// TIA Portal project "Lagerregal_5" (V20) (continued)

   IF #"PTRIG_MDB_Z-Neg".Q THEN
       "HMI_Schnittstelle".Kraene.Kran_1.Kran_Pos."Z-Soll" -= UINT_TO_INT("HMI_Schnittstelle".HMI.Inkrement);
   END_IF;
END_REGION
END_FUNCTION_BLOCK

FUNCTION_BLOCK "Ein_HMI"   // FB10, FBD
{ S7_Optimized_Access := 'TRUE' }
VERSION : 0.1
BEGIN
END_FUNCTION_BLOCK

FUNCTION "Meldungen" : Void   // FC10, SCL
{ S7_Optimized_Access := 'TRUE' }
VERSION : 0.1
BEGIN
   // Slice Zugriff programmieren
   // d.h. wir können auf die Einzelbits einer Ganzzahlvariable (INT, DINT, etc.)
   // bzw. einer Bitfolge (Byte, Word, etc.) zugreifen.

   // Bits:        Variable.%X0
   // Bytes:       Variable.%B0
   // Word:        Variable.%W0
   // DWord:       Variable.%D0


   "HMI_Schnittstelle".Bitmeldungen.%X0 := "HMI_Schnittstelle".Eingaenge.S2;
   "HMI_Schnittstelle".Bitmeldungen.%X1 := "HMI_Schnittstelle".Eingaenge.S1;
   "HMI_Schnittstelle".Bitmeldungen.%X2 := "HMI_Schnittstelle".Betriebsart.Hand;
   "HMI_Schnittstelle".Bitmeldungen.%X3 := "HMI_Schnittstelle".Betriebsart.Automatik;
END_FUNCTION

// folder: Kransteuerung

FUNCTION_BLOCK "FC_Kran_beladen"   // FB25, FBD
{ S7_Optimized_Access := 'TRUE' }
VERSION : 0.1
   VAR_INPUT
      "eKran_Z-Ist" : Int;
      eSchrittnummer : Int;
   END_VAR
   VAR_OUTPUT
      aGabel : Bool;
      aBeladen : Bool;
      "aKran_Z-Soll" : Int;
   END_VAR
   VAR
      PTRIG_Schritt2 : Bool;
   END_VAR
   VAR_TEMP   // added for the SCL form of the ladder/FBD networks
      _w1 : Bool;
      _w2 : Bool;
   END_VAR
BEGIN

REGION Network 1: Gabel zur Seite ausfahren
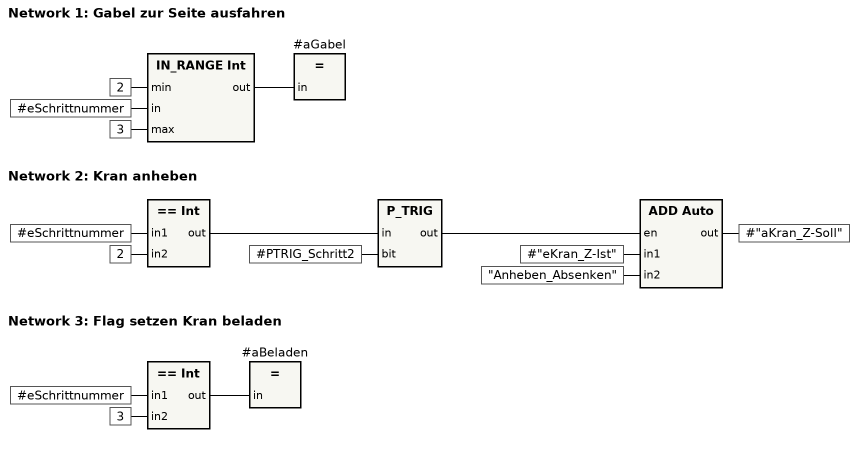
   #aGabel := (2 <= #eSchrittnummer) AND (#eSchrittnummer <= 3);
END_REGION

REGION Network 2: Kran anheben
   #_w1 := #eSchrittnummer = 2;
   #_w2 := #_w1 AND NOT #PTRIG_Schritt2;   // rising edge
   #PTRIG_Schritt2 := #_w1;
   IF #_w2 THEN #"aKran_Z-Soll" := #"eKran_Z-Ist" + "Anheben_Absenken"; END_IF;
END_REGION

REGION Network 3: Flag setzen Kran beladen
   #aBeladen := #eSchrittnummer = 3;
END_REGION
END_FUNCTION_BLOCK

FUNCTION_BLOCK "FC_Kran_entladen"   // FB26, FBD
{ S7_Optimized_Access := 'TRUE' }
VERSION : 0.1
   VAR_INPUT
      "eKran_Z-Ist" : Int;
      eSchrittnummer : Int;
   END_VAR
   VAR_OUTPUT
      aGabel : Bool;
      aBeladen : Bool;
      "aKran_Z-Soll" : Int;
   END_VAR
   VAR
      PTRIG_Schritt2 : Bool;
   END_VAR
   VAR_TEMP   // added for the SCL form of the ladder/FBD networks
      _w1 : Bool;
      _w2 : Bool;
   END_VAR
BEGIN

REGION Network 1: Gabel zur Seite ausfahren
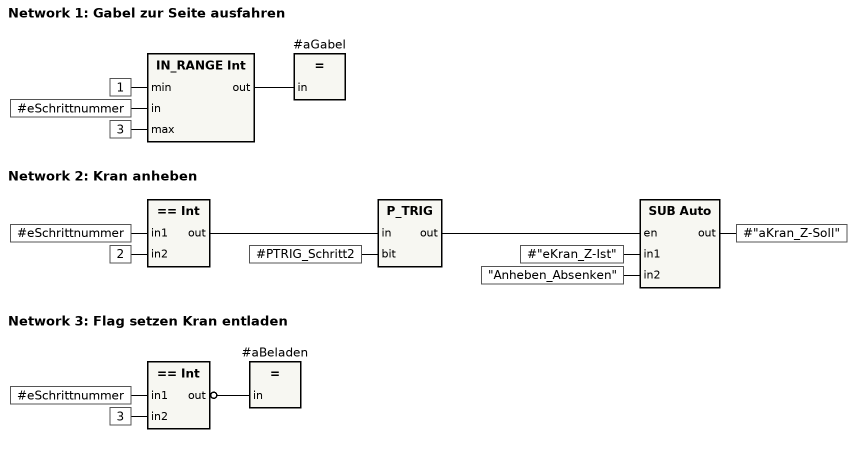
   #aGabel := (1 <= #eSchrittnummer) AND (#eSchrittnummer <= 3);
END_REGION

REGION Network 2: Kran anheben
   #_w1 := #eSchrittnummer = 2;
   #_w2 := #_w1 AND NOT #PTRIG_Schritt2;   // rising edge
   #PTRIG_Schritt2 := #_w1;
   IF #_w2 THEN #"aKran_Z-Soll" := #"eKran_Z-Ist" - "Anheben_Absenken"; END_IF;
END_REGION

REGION Network 3: Flag setzen Kran entladen
   #aBeladen := NOT (#eSchrittnummer = 3);
END_REGION
END_FUNCTION_BLOCK

FUNCTION_BLOCK "Ein_Kran"   // FB30, FBD
{ S7_Optimized_Access := 'TRUE' }
VERSION : 0.1
   VAR
      NTRIG_MDB_1B2 : F_TRIG;
      NTRIG_MDB_2B2 : F_TRIG;
      NTRIG_MDB_5B1 : F_TRIG;
   END_VAR
BEGIN

REGION Network 1 (SCL): Sensoren Kran_1
   "HMI_Schnittstelle".Eingaenge."6B1" := "6B1";
   "HMI_Schnittstelle".Eingaenge."6B2" := "6B2";
   "HMI_Schnittstelle".Eingaenge."6B3" := "6B3";
END_REGION

REGION Network 2: Kran_1 Position einlesen
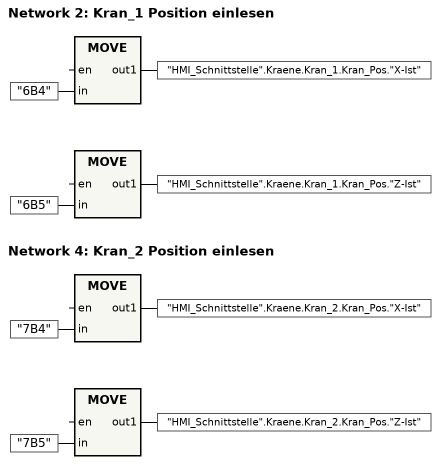
   "HMI_Schnittstelle".Kraene.Kran_1.Kran_Pos."X-Ist" := "6B4";
   "HMI_Schnittstelle".Kraene.Kran_1.Kran_Pos."Z-Ist" := "6B5";
END_REGION

REGION Network 3 (SCL): Sensoren Kran_2
   "HMI_Schnittstelle".Eingaenge."7B1" := "7B1";
   "HMI_Schnittstelle".Eingaenge."7B2" := "7B2";
   "HMI_Schnittstelle".Eingaenge."7B3" := "7B3";
END_REGION

REGION Network 4: Kran_2 Position einlesen
   "HMI_Schnittstelle".Kraene.Kran_2.Kran_Pos."X-Ist" := "7B4";
   "HMI_Schnittstelle".Kraene.Kran_2.Kran_Pos."Z-Ist" := "7B5";
END_REGION
END_FUNCTION_BLOCK

FUNCTION_BLOCK "Prog_Automatik_einlagern"   // FB50, FBD
{ S7_Optimized_Access := 'TRUE' }
VERSION : 0.1
   VAR
      MDB_Schrittkette_einlagern : "Prog_Schrittkette";
      FTRIG_Palette_eingelagert : F_TRIG;
   END_VAR
   VAR_TEMP
      tmpPalette_abgelegt : Int;
      tmpFaecher_durchlaufen : Int;
   END_VAR
BEGIN

REGION Network 1 (SCL): Lagerplatz frei
   IF "HMI_Schnittstelle".Anlagendaten.Fach > 0 AND "HMI_Schnittstelle".Anlagendaten.Fach < 55 THEN
       "HMI_Schnittstelle".Anlagendaten.Regalplatz_frei := "Warenlager".Lager["HMI_Schnittstelle".Anlagendaten.Fach].Bauteil = 0;

       IF NOT "HMI_Schnittstelle".Anlagendaten.Regalplatz_frei AND "HMI_Schnittstelle".Anlagendaten.Fach < 54 THEN
           // Zähle das Fach hoch, wenn das aktuell Fach belegt ist.
           "HMI_Schnittstelle".Anlagendaten.Fach += 1;
       END_IF;
   ELSE
       "HMI_Schnittstelle".Anlagendaten.Regalplatz_frei := FALSE;
   END_IF;


   // Verhindere Endlos-Schleife
   IF #tmpFaecher_durchlaufen = 2 AND NOT "HMI_Schnittstelle".Anlagendaten.Regalplatz_frei THEN
       "HMI_Schnittstelle".Anlagendaten.Fach := 0;
       "HMI_Schnittstelle".Betriebsart.Automatik := FALSE;
   END_IF;
END_REGION

REGION Network 2: Palette abgelegt
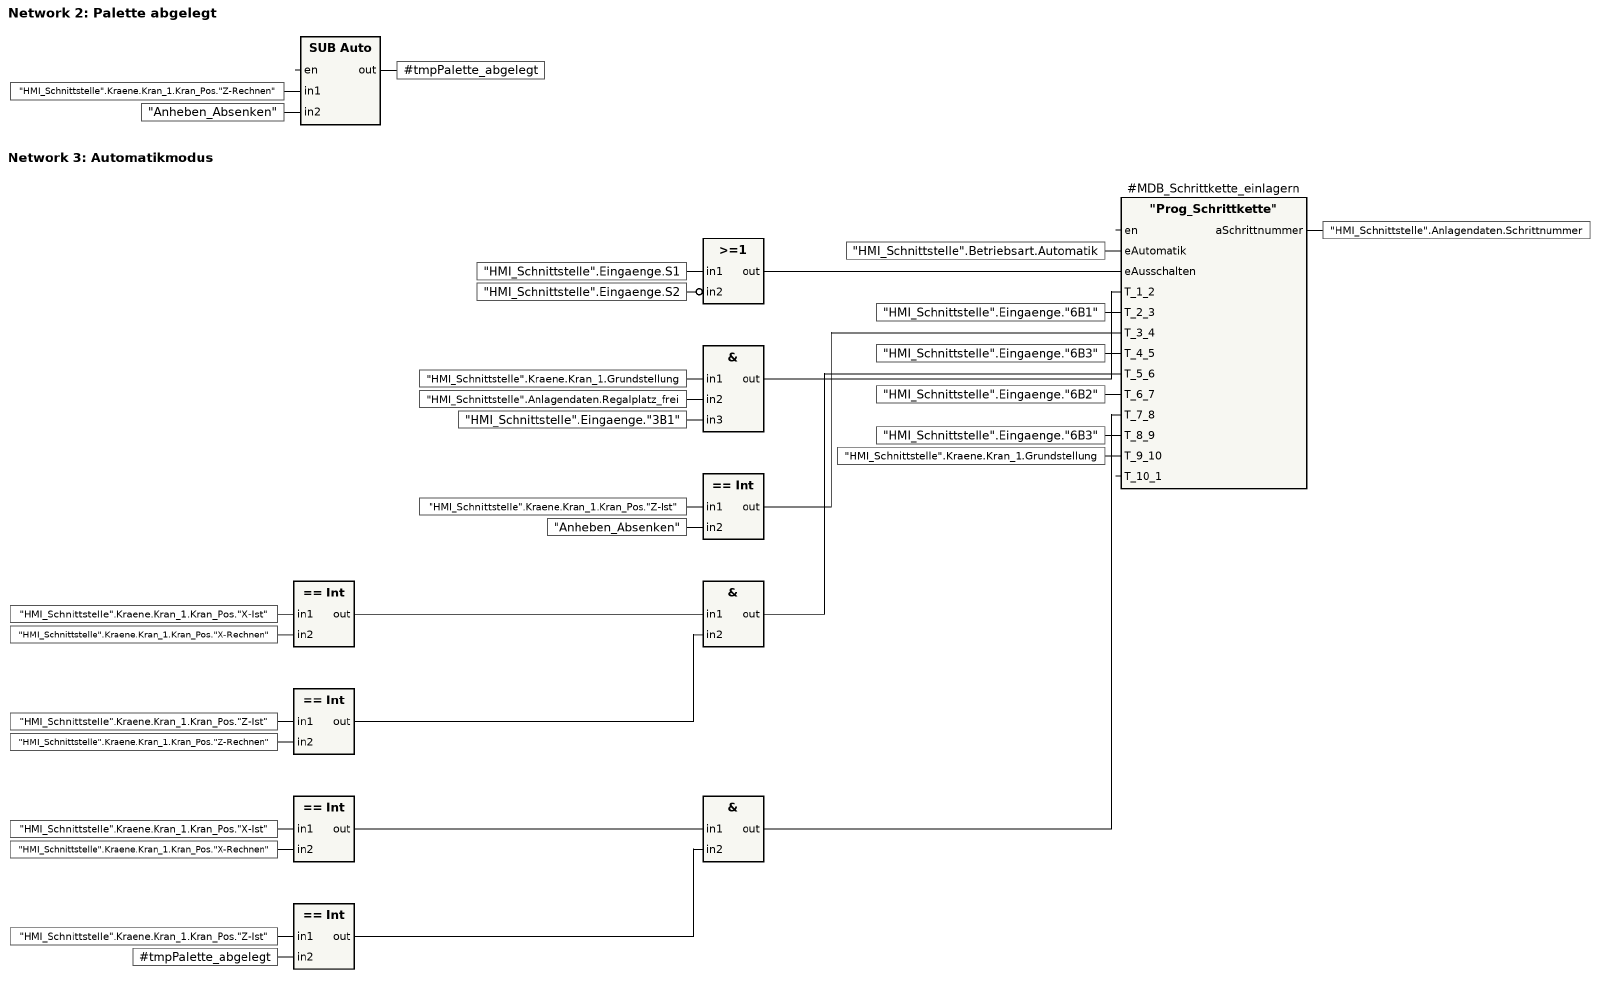
   #tmpPalette_abgelegt := "HMI_Schnittstelle".Kraene.Kran_1.Kran_Pos."Z-Rechnen" - "Anheben_Absenken";
END_REGION

REGION Network 3: Automatikmodus
   #MDB_Schrittkette_einlagern(eAutomatik := "HMI_Schnittstelle".Betriebsart.Automatik,   // "Prog_Schrittkette"
                           eAusschalten := "HMI_Schnittstelle".Eingaenge.S1 OR NOT "HMI_Schnittstelle".Eingaenge.S2,
                           T_1_2 := "HMI_Schnittstelle".Kraene.Kran_1.Grundstellung AND "HMI_Schnittstelle".Anlagendaten.Regalplatz_frei AND "HMI_Schnittstelle".Eingaenge."3B1",
                           T_2_3 := "HMI_Schnittstelle".Eingaenge."6B1",
                           T_3_4 := "HMI_Schnittstelle".Kraene.Kran_1.Kran_Pos."Z-Ist" = "Anheben_Absenken",
                           T_4_5 := "HMI_Schnittstelle".Eingaenge."6B3",
                           T_5_6 := ("HMI_Schnittstelle".Kraene.Kran_1.Kran_Pos."X-Ist" = "HMI_Schnittstelle".Kraene.Kran_1.Kran_Pos."X-Rechnen") AND ("HMI_Schnittstelle".Kraene.Kran_1.Kran_Pos."Z-Ist" = "HMI_Schnittstelle".Kraene.Kran_1.Kran_Pos."Z-Rechnen"),
                           T_6_7 := "HMI_Schnittstelle".Eingaenge."6B2",
                           T_7_8 := ("HMI_Schnittstelle".Kraene.Kran_1.Kran_Pos."X-Ist" = "HMI_Schnittstelle".Kraene.Kran_1.Kran_Pos."X-Rechnen") AND ("HMI_Schnittstelle".Kraene.Kran_1.Kran_Pos."Z-Ist" = #tmpPalette_abgelegt),
                           T_8_9 := "HMI_Schnittstelle".Eingaenge."6B3",
                           T_9_10 := "HMI_Schnittstelle".Kraene.Kran_1.Grundstellung,
                           aSchrittnummer => "HMI_Schnittstelle".Anlagendaten.Schrittnummer);
END_REGION

REGION Network 4 (SCL): Fachnummer erhöhen
   #FTRIG_Palette_eingelagert(CLK := "HMI_Schnittstelle".Anlagendaten.Schrittnummer = 7);


   // Wenn die Palette eingelagert wurde, ...
   IF #FTRIG_Palette_eingelagert.Q THEN
       // ... schreibe die Info über das Bauteil ins Array.
       "Warenlager".Lager["HMI_Schnittstelle".Anlagendaten.Fach].Bauteil := "HMI_Schnittstelle".Anlagendaten.Bauteil;

       // Zähle das Fach hoch und setze das aktuelle Bauteil zurück.
       "HMI_Schnittstelle".Anlagendaten.Fach += 1;
       "HMI_Schnittstelle".Anlagendaten.Bauteil := 0;
   END_IF;

   IF "HMI_Schnittstelle".Anlagendaten.Fach = 54 THEN
       // Setze das Fach 1, wenn am Ende angekommen.
       "HMI_Schnittstelle".Anlagendaten.Fach := 1;
       #tmpFaecher_durchlaufen += 1;
   END_IF;
END_REGION
END_FUNCTION_BLOCK

FUNCTION "Aus_Kran" : Void   // FC30, FBD
{ S7_Optimized_Access := 'TRUE' }
VERSION : 0.1
BEGIN

REGION Network 1 (SCL): Kräne Gabelsteuerung
   "6M1" := "HMI_Schnittstelle".Ausgaenge."6M1";
   "6M2" := "HMI_Schnittstelle".Ausgaenge."6M2";

   "7M1" := "HMI_Schnittstelle".Ausgaenge."7M1";
   "7M2" := "HMI_Schnittstelle".Ausgaenge."7M2";
END_REGION
END_FUNCTION

FUNCTION "FC_Kran_Grundstellung" : Void   // FC31, FBD
{ S7_Optimized_Access := 'TRUE' }
VERSION : 0.1
   VAR_INPUT
      "X-Ist" : Int;
      "Z-Ist" : Int;
      Gabel_mitte : Bool;
   END_VAR
   VAR_OUTPUT
      Heimposition : Bool;
      Grundstellung : Bool;
   END_VAR
BEGIN

REGION Network 1
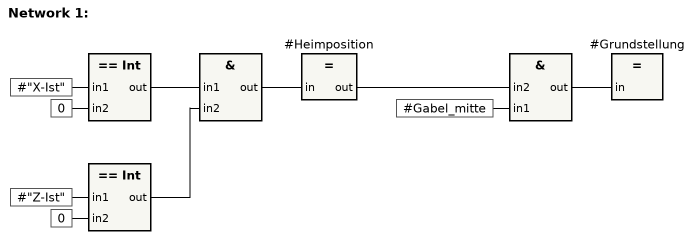
   #Heimposition := (#"X-Ist" = 0) AND (#"Z-Ist" = 0);
   #Grundstellung := #Heimposition AND #Gabel_mitte;
END_REGION
END_FUNCTION

FUNCTION "Staplersteuerung" : Void   // FC70, FBD
{ S7_Optimized_Access := 'TRUE' }
VERSION : 0.1
BEGIN

REGION Network 1: Sollposition X
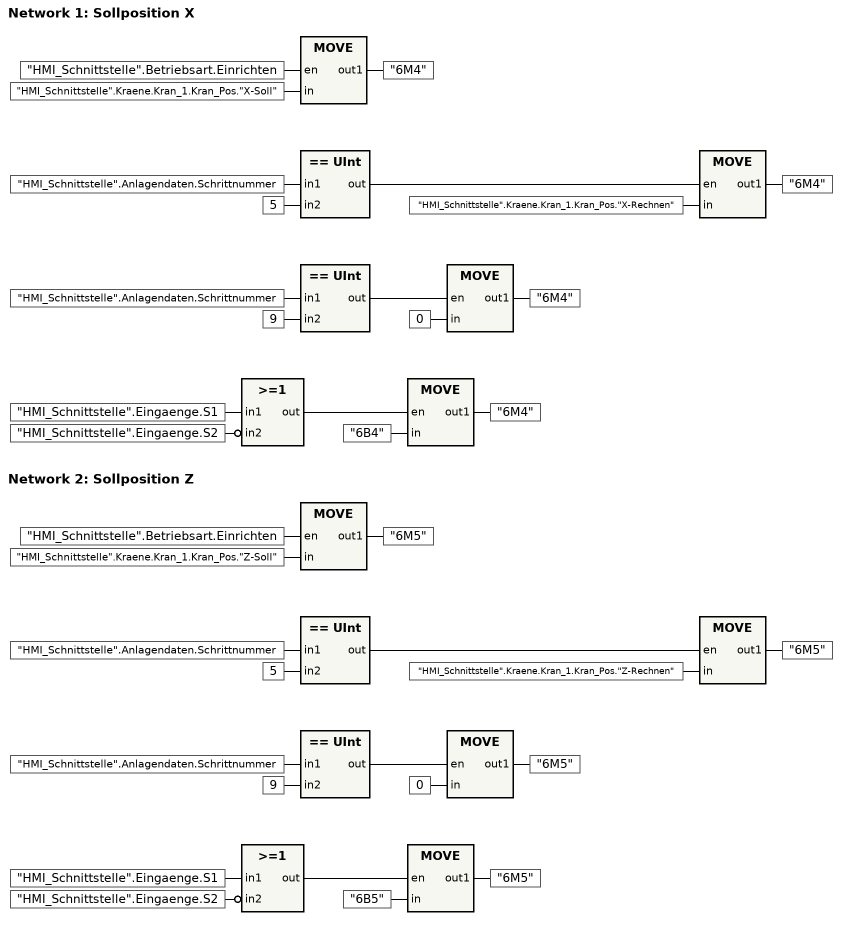
   IF "HMI_Schnittstelle".Betriebsart.Einrichten THEN
       "6M4" := "HMI_Schnittstelle".Kraene.Kran_1.Kran_Pos."X-Soll";
   END_IF;
   IF "HMI_Schnittstelle".Anlagendaten.Schrittnummer = 5 THEN
       "6M4" := "HMI_Schnittstelle".Kraene.Kran_1.Kran_Pos."X-Rechnen";
   END_IF;
   IF "HMI_Schnittstelle".Anlagendaten.Schrittnummer = 9 THEN "6M4" := 0; END_IF;
   IF "HMI_Schnittstelle".Eingaenge.S1 OR NOT "HMI_Schnittstelle".Eingaenge.S2 THEN "6M4" := "6B4"; END_IF;
END_REGION

REGION Network 2: Sollposition Z
   IF "HMI_Schnittstelle".Betriebsart.Einrichten THEN
       "6M5" := "HMI_Schnittstelle".Kraene.Kran_1.Kran_Pos."Z-Soll";
   END_IF;
   IF "HMI_Schnittstelle".Anlagendaten.Schrittnummer = 5 THEN
       "6M5" := "HMI_Schnittstelle".Kraene.Kran_1.Kran_Pos."Z-Rechnen";
   END_IF;
   IF "HMI_Schnittstelle".Anlagendaten.Schrittnummer = 9 THEN "6M5" := 0; END_IF;
   IF "HMI_Schnittstelle".Eingaenge.S1 OR NOT "HMI_Schnittstelle".Eingaenge.S2 THEN "6M5" := "6B5"; END_IF;
END_REGION

REGION Network 3 (SCL): Z-Achse Kran_1 Soll-Pos
   (*
   IF NOT "HMI_Schnittstelle".Eingaenge.S2 OR "HMI_Schnittstelle".Eingaenge.S1 THEN
       ;
   *)

   // Einrichtbetrieb
   IF "HMI_Schnittstelle".Betriebsart.Einrichten THEN
       "6M5" := "HMI_Schnittstelle".Kraene.Kran_1.Kran_Pos."Z-Soll";

   // Automatikbetrieb    
   ELSIF "HMI_Schnittstelle".Anlagendaten.Schrittnummer = 3 THEN
       // Palette aus Grundstellung anheben
       "6M5" := "Anheben_Absenken" + 2;
   ELSIF "HMI_Schnittstelle".Anlagendaten.Schrittnummer = 5 THEN
       //Fach mit Nummer anfahren
       "6M5" := "HMI_Schnittstelle".Kraene.Kran_1.Kran_Pos."Z-Rechnen";
   ELSIF "HMI_Schnittstelle".Anlagendaten.Schrittnummer = 7 THEN
       // Palette in Regal einlagern
       "6M5" := "HMI_Schnittstelle".Kraene.Kran_1.Kran_Pos."Z-Rechnen" - "Anheben_Absenken";
   ELSIF "HMI_Schnittstelle".Anlagendaten.Schrittnummer = 9 THEN
       // Stapler in Grundstellung
       "6M5" := 0;
   END_IF;
END_REGION

REGION Network 4 (SCL): Gabel links ausfahren
   "HMI_Schnittstelle".Ausgaenge."6M1" := "HMI_Schnittstelle".Anlagendaten.Schrittnummer = 2
                                       OR "HMI_Schnittstelle".Anlagendaten.Schrittnummer = 3;
END_REGION

REGION Network 5 (SCL): Gabel rechts ausfahren
   "HMI_Schnittstelle".Ausgaenge."6M2" := "HMI_Schnittstelle".Anlagendaten.Schrittnummer = 6
                                       OR "HMI_Schnittstelle".Anlagendaten.Schrittnummer = 7;
END_REGION
END_FUNCTION

ORGANIZATION_BLOCK "Main_einlagern"   // OB123, FBD, ProgramCycle
TITLE = "Main Program Sweep (Cycle)"
{ S7_Optimized_Access := 'TRUE' }
VERSION : 0.1
   VAR_INPUT
      Initial_Call : Bool;   // Initial call of this OB
      Remanence : Bool;   // =True, if remanent data are available
   END_VAR
BEGIN

REGION Network 1: Test ob Kran in Grundstellung ist
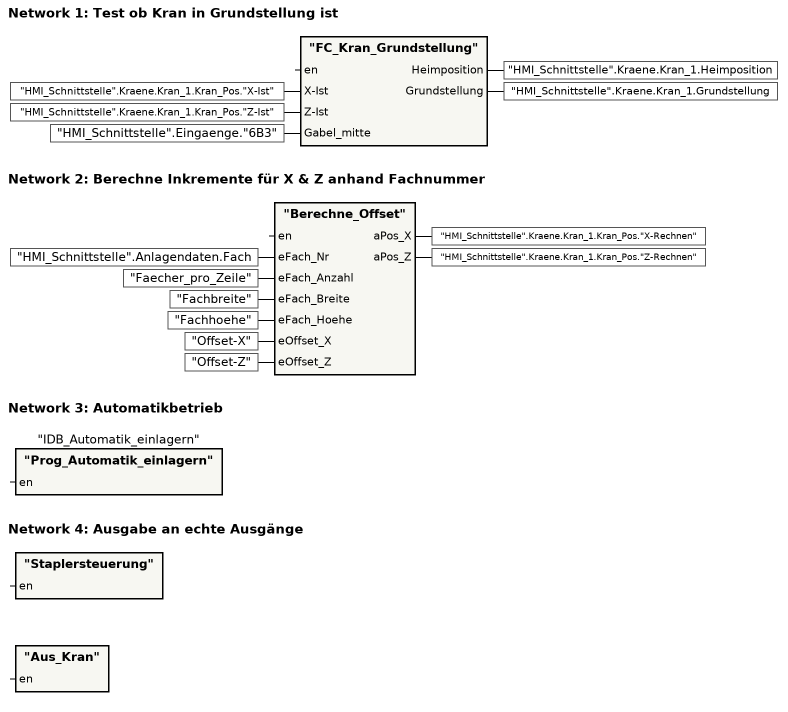
   "FC_Kran_Grundstellung"("X-Ist" := "HMI_Schnittstelle".Kraene.Kran_1.Kran_Pos."X-Ist",
                           "Z-Ist" := "HMI_Schnittstelle".Kraene.Kran_1.Kran_Pos."Z-Ist",
                           Gabel_mitte := "HMI_Schnittstelle".Eingaenge."6B3",
                           Heimposition => "HMI_Schnittstelle".Kraene.Kran_1.Heimposition,
                           Grundstellung => "HMI_Schnittstelle".Kraene.Kran_1.Grundstellung);
END_REGION

REGION Network 2: Berechne Inkremente für X & Z anhand Fachnummer
   "Berechne_Offset"(eFach_Nr := "HMI_Schnittstelle".Anlagendaten.Fach,
                     eFach_Anzahl := "Faecher_pro_Zeile",
                     eFach_Breite := "Fachbreite",
                     eFach_Hoehe := "Fachhoehe",
                     eOffset_X := "Offset-X",
                     eOffset_Z := "Offset-Z",
                     aPos_X => "HMI_Schnittstelle".Kraene.Kran_1.Kran_Pos."X-Rechnen",
                     aPos_Z => "HMI_Schnittstelle".Kraene.Kran_1.Kran_Pos."Z-Rechnen");
END_REGION

REGION Network 3: Automatikbetrieb
   "IDB_Automatik_einlagern"();   // "Prog_Automatik_einlagern"
END_REGION

REGION Network 4: Ausgabe an echte Ausgänge
   "Staplersteuerung"();
   "Aus_Kran"();
END_REGION
END_ORGANIZATION_BLOCK

(* ===== HMI "HMI_RT_1" =====
system functions are stored by id; their names below are inferred from use
connection "HMI_Verbindung_1": ETHERNET, S7_1500_OMS

HMI tags "Standard-Variablentabelle"
   "HMI_Schnittstelle_Kraene_Kran_1_Z-Soll" : Int = PLC HMI_Schnittstelle.Kraene.Kran_1.Kran_Pos.Z-Soll, 100 ms
   "HMI_Schnittstelle_Kraene_Kran_1_X-Soll" : Int = PLC HMI_Schnittstelle.Kraene.Kran_1.Kran_Pos.X-Soll, 100 ms
   "HMI_Schnittstelle_Kraene_Kran_1_X-Ist" : Int = PLC HMI_Schnittstelle.Kraene.Kran_1.Kran_Pos.X-Ist, 100 ms
   "HMI_Schnittstelle_Kraene_Kran_1_Z-Ist" : Int = PLC HMI_Schnittstelle.Kraene.Kran_1.Kran_Pos.Z-Ist, 100 ms
   "HMI_Schnittstelle_HMI_X-Neg" : Bool = PLC HMI_Schnittstelle.HMI.X-Neg, 1 s
   "HMI_Schnittstelle_HMI_X-Pos" : Bool = PLC HMI_Schnittstelle.HMI.X-Pos, 1 s
   "HMI_Schnittstelle_HMI_Z-Neg" : Bool = PLC HMI_Schnittstelle.HMI.Z-Neg, 1 s
   "HMI_Schnittstelle_HMI_Z-Pos" : Bool = PLC HMI_Schnittstelle.HMI.Z-Pos, 1 s
   "HMI_Schnittstelle_HMI_Inkrement" : UInt = PLC HMI_Schnittstelle.HMI.Inkrement, 1 s
   "Clock_1Hz" : Bool = PLC Clock_1Hz AT %M0.5, 100 ms
   "HMI_Schnittstelle_Fach" : Int = PLC HMI_Schnittstelle.Anlagendaten.Fach, 500 ms
   "HMI_Schnittstelle_Fach_ansteuern" : Bool = PLC HMI_Schnittstelle.Anlagendaten.Fach_ansteuern, 1 s
   "Warenlager_Lager{1}_Flags_Belegt" : Bool = PLC Warenlager.Lager[1].Flags.Belegt, 1 s
   "Warenlager_Lager{1}_Flags_In_Benutzung" : Bool = PLC Warenlager.Lager[1].Flags.In_Benutzung, 1 s
   "HMI_Schnittstelle_Anlagendaten_Schrittnummer" : UInt = PLC HMI_Schnittstelle.Anlagendaten.Schrittnummer, 100 ms
   "HMI_Schnittstelle_Bitmeldungen" : Word = PLC HMI_Schnittstelle.Bitmeldungen, 1 s
   "HMI_Schnittstelle_Betriebsart_Einrichten" : Bool = PLC HMI_Schnittstelle.Betriebsart.Einrichten, 1 s
   "HMI_Schnittstelle_Betriebsart_Automatik" : Bool = PLC HMI_Schnittstelle.Betriebsart.Automatik, 1 s
   "HMI_Schnittstelle_Betriebsart_Hand" : Bool = PLC HMI_Schnittstelle.Betriebsart.Hand, 1 s

HMI tags "Interne_Variablen"
   "Bildnummer" : Int, internal
   "Benutzername" : WString[254], internal
   "Anz_Anmeldungen" : UDInt, internal

discrete alarms
   1: 'Hauptschalter wurde eingeschaltet', class Warnings, trigger "HMI_Schnittstelle_Bitmeldungen" bit 0
   2: 'Not-Halt wurde betätigt', class Errors, trigger "HMI_Schnittstelle_Bitmeldungen" bit 1
   3: 'Handbetrieb wurde aktiviert', class Warnings, trigger "HMI_Schnittstelle_Bitmeldungen" bit 2
   4: 'Automatik wurde gestartet', class Warnings, trigger "HMI_Schnittstelle_Bitmeldungen" bit 3

analog alarms
   1: 'Stapler hat Palette aufgenommen', class Anzeigen, trigger "HMI_Schnittstelle_Anlagendaten_Schrittnummer"
   2: 'Stapler fährt zu Fach', class Anzeigen, trigger "HMI_Schnittstelle_Anlagendaten_Schrittnummer"
   3: 'Stapler hat Palette abgelegt', class Anzeigen, trigger "HMI_Schnittstelle_Anlagendaten_Schrittnummer"
   4: 'Benutzername', class Anzeigen, trigger "Anz_Anmeldungen"

text list "Liste_Bilder": 0..1 'Bitte Bild auswählen'; 1 'Startbild'; 2 'Betriebsart'; 3 'Handbetrieb'; 4 ''; 5 'Einrichtbetrieb'; 6 'Statistik'; 7 ''; 8 'Meldungen'; 9 'Diagnose'; 10 'Benutzerverwaltung'

screen "01_0_Lageransicht" 800x420, template "Menüleiste"
   on GenerateScreen: SetTag("Bildnummer", 1)
   Button "Schaltfläche_4" at 10,438 size 96x32; TextOff 'Teachen'
      on Press: ActivateScreen("05_Einrichtbetrieb", 0)
   Rectangle "Rechteck_1" at 650,280 size 50x50
      Appearance <- "Warenlager_Lager{1}_Flags_Belegt"
   TextField "Textfeld_1" at 650,280 size 50x50; Text '1'
      Appearance <- "Warenlager_Lager{1}_Flags_In_Benutzung"
   GraphicView "Grafikanzeige_1" at 275,170 size 50x50; Picture "Palette"
      DiagonalMovement <- "HMI_Schnittstelle_Kraene_Kran_1_X-Ist"
   TextField "Textfeld_2" at 89,10 size 163x23; Text 'Stapler einlagern'

screen "05_Einrichtbetrieb" 800x420, template "Menüleiste"
   on GenerateScreen: SetTag("Bildnummer", 5)
   on ClearScreen: function_f23ef4c9()
   Button "Schaltfläche_1" at 694,10 size 96x32; TextOff 'Zurück'
      on Press: function_efd93a16()
   TextField "Textfeld_1" at 308,10 size 184x23; Text 'Kalibrierungsmodus'
   Slider "Schieberegler_2" at 113,300 size 230x50; Caption 'Breite'
      ProcessValue <- "HMI_Schnittstelle_Kraene_Kran_1_X-Soll"
   IOField "EA-Feld_8" at 370,67 size 96x32; FormatPattern 99999
      ProcessValue <- "HMI_Schnittstelle_Kraene_Kran_1_X-Ist"
   IOField "EA-Feld_9" at 485,68 size 96x32; FormatPattern 99999
      ProcessValue <- "HMI_Schnittstelle_Kraene_Kran_1_Z-Ist"
   Slider "Schieberegler_1" at 10,37 size 50x230; Caption 'Höhe'
      ProcessValue <- "HMI_Schnittstelle_Kraene_Kran_1_Z-Soll"
   Button "Schaltfläche_5" at 345,300 size 25x50; TextOff '-'
      on Press: function_b14e0dd5("HMI_Schnittstelle_HMI_X-Neg", 0)
      Appearance <- "HMI_Schnittstelle_HMI_X-Neg"
   IOField "EA-Feld_7" at 10,300 size 70x50; FormatPattern 99999
      ProcessValue <- "HMI_Schnittstelle_HMI_Inkrement"
   Button "Schaltfläche_7" at 10,269 size 50x25; TextOff '-'
      on Press: function_b14e0dd5("HMI_Schnittstelle_HMI_Z-Neg", 0)
      Appearance <- "HMI_Schnittstelle_HMI_Z-Neg"
   Button "Schaltfläche_8" at 10,10 size 50x25; TextOff '+'
      on Press: function_b14e0dd5("HMI_Schnittstelle_HMI_Z-Pos", 0)
      Appearance <- "HMI_Schnittstelle_HMI_Z-Pos"
   Button "Schaltfläche_6" at 86,300 size 25x50; TextOff '+'
      on Press: function_b14e0dd5("HMI_Schnittstelle_HMI_X-Pos", 0)
      Appearance <- "HMI_Schnittstelle_HMI_X-Pos"
   TextField "Textfeld_2" at 370,42 size 111x23; Text 'Ist-X-Achse'
   TextField "Textfeld_3" at 485,42 size 110x23; Text 'Ist-Z-Achse'
   TextField "Textfeld_4" at 370,103 size 88x23; Text 'Fach-Nr.:'
   IOField "EA-Feld_1" at 370,128 size 96x32; FormatPattern 99
      ProcessValue <- "HMI_Schnittstelle_Fach"
   Button "Schaltfläche_2" at 485,128 size 96x32; TextOff 'Testen'
      on Press: function_b14e0dd5("HMI_Schnittstelle_Fach_ansteuern", 0)

screen "01_1_Detailansicht" 800x420, template "Menüleiste"
   Button "Schaltfläche_1" at 694,10 size 96x32; TextOff 'Zurück'
      on Press: function_efd93a16()

Template "Menüleiste" 800x420
   Button "Vorlage_Schaltfläche_1" at 0,360 size 80x60; TextOff 'HOME'; PictureOff "Grafik_2"; PictureOn "Grafik_2"
      Appearance <- "Bildnummer"
      on Press: ActivateScreen("01_0_Lageransicht", 0)
   Button "Vorlage_Schaltfläche_2" at 80,360 size 80x60; TextOff 'BETRIEB'; PictureOff "Grafik_8"; PictureOn "Grafik_8"
      Appearance <- "Bildnummer"
      on Press: ActivateScreen("02_Betriebsart", 0)
   Button "Vorlage_Schaltfläche_3" at 160,360 size 80x60; TextOff 'HAND'; PictureOff "Grafik_7"; PictureOn "Grafik_7"
      Appearance <- "Bildnummer"
      on Press: ActivateScreen("03_Bild", 0)
   Button "Vorlage_Schaltfläche_4" at 240,360 size 80x60; TextOff 'Text'
      Appearance <- "Bildnummer"
      on Press: ActivateScreen("04_Bild", 0)
   Button "Vorlage_Schaltfläche_5" at 320,360 size 80x60; TextOff 'TEACH'; PictureOn "Grafik_3"; PictureOff "Grafik_3"; Authorization "Einstellen"
      Appearance <- "Bildnummer"
      on Press: SetTag("HMI_Schnittstelle_Betriebsart_Einrichten", 1); SetTag("HMI_Schnittstelle_Betriebsart_Automatik", 0); SetTag("HMI_Schnittstelle_Betriebsart_Hand", 0); ActivateScreen("05_Einrichtbetrieb", 0)
   Button "Vorlage_Schaltfläche_6" at 400,360 size 80x60; TextOff 'STATS'; PictureOff "Grafik_4"; PictureOn "Grafik_4"
      Appearance <- "Bildnummer"
      on Press: ActivateScreen("06_Statistik", 0)
   Button "Vorlage_Schaltfläche_7" at 480,360 size 80x60; TextOff 'Text'
      Appearance <- "Bildnummer"
      on Press: ActivateScreen("07_Bild", 0)
   Button "Vorlage_Schaltfläche_8" at 560,360 size 80x60; TextOff 'FEHLER'; PictureOff "Grafik_6"; PictureOn "Grafik_6"
      Appearance <- "Bildnummer"
      on Press: ActivateScreen("08_0_Meldungen", 0)
   Button "Vorlage_Schaltfläche_9" at 640,360 size 80x60; TextOff 'DIAG'; PictureOff "Grafik_9"; PictureOn "Grafik_9"
      Appearance <- "Bildnummer"
      on Press: ActivateScreen("09_Diagnose", 0)
   Button "Vorlage_Schaltfläche_10" at 720,360 size 80x60; TextOff 'NUTZER'; PictureOff "Grafik_10"; PictureOn "Grafik_10"
      Appearance <- "Bildnummer"
      on Press: ActivateScreen("10_Benutzer", 0)

screen "02_Betriebsart" 800x420, template "Menüleiste"
   on GenerateScreen: SetTag("Bildnummer", 2)

screen "03_Bild" 800x420, template "Menüleiste"
   on GenerateScreen: SetTag("Bildnummer", 3)

screen "04_Bild" 800x420, template "Menüleiste"
   on GenerateScreen: SetTag("Bildnummer", 4)

screen "06_Statistik" 800x420, template "Menüleiste"
   on GenerateScreen: SetTag("Bildnummer", 6)
   TrendView "Kurvenanzeige_1" at 10,10 size 780x340

screen "07_Bild" 800x420, template "Menüleiste"
   on GenerateScreen: SetTag("Bildnummer", 7)

screen "08_0_Meldungen" 800x420, template "Menüleiste"
   on GenerateScreen: SetTag("Bildnummer", 8)
   AlarmView "Meldeanzeige_1" at 10,50 size 780x300
   TextField "Textfeld_1" at 10,10 size 103x23; Text 'Meldungen'
   Button "Schaltfläche_1" at 598,11 size 192x32; TextOff '08_1_Meldepuffer'
      on Click: ActivateScreen("08_1_Meldepuffer", 0)

screen "09_Diagnose" 800x420, template "Menüleiste"
   on GenerateScreen: SetTag("Bildnummer", 9)
   SysDiagControl "System-Diagnoseanzeige_1" at 10,10 size 780x340

screen "10_Benutzer" 800x420, template "Menüleiste"
   on GenerateScreen: SetTag("Bildnummer", 10)
   UserView "Benutzeranzeige_1" at 10,10 size 780x340

screen "08_1_Meldepuffer" 800x420, template "Menüleiste"
   on GenerateScreen: SetTag("Bildnummer", 8)
   AlarmView "Meldeanzeige_1" at 10,50 size 780x300
   TextField "Textfeld_1" at 10,10 size 114x23; Text 'Meldepuffer'
   Button "Schaltfläche_1" at 598,10 size 192x32; TextOff '08_0_Meldungen'
      on Click: ActivateScreen("08_0_Meldungen", 0)

scheduled task "Anmeldung"
   on Action: function_f41c6f6c("Benutzername"); function_dd21b452("Anz_Anmeldungen", 1)
*)